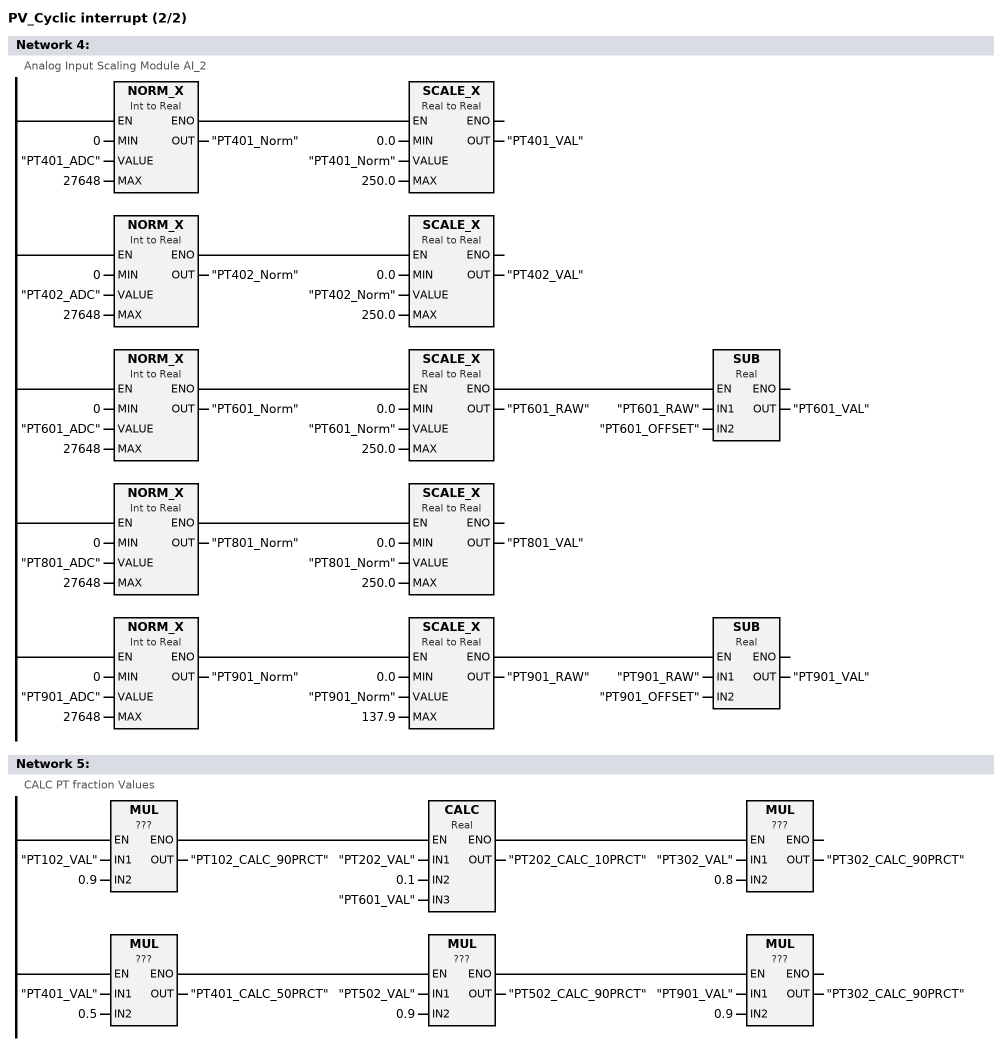
   RUNG wire#powerrail
      { S7_Templates := "[SrcType := Int, DestType := Real]" } Normalize(min := 0, value := "PT401_ADC", max := 27648, out => "PT401_Norm")
      { S7_Templates := "[SrcType := Real, DestType := Real]" } Scale(min := 0.0, value := "PT401_Norm", max := 250.0, out => "PT401_VAL")
   END_RUNG
   RUNG wire#powerrail
      { S7_Templates := "[SrcType := Int, DestType := Real]" } Normalize(min := 0, value := "PT402_ADC", max := 27648, out => "PT402_Norm")
      { S7_Templates := "[SrcType := Real, DestType := Real]" } Scale(min := 0.0, value := "PT402_Norm", max := 250.0, out => "PT402_VAL")
   END_RUNG
   RUNG wire#powerrail
      { S7_Templates := "[SrcType := Int, DestType := Real]" } Normalize(min := 0, value := "PT601_ADC", max := 27648, out => "PT601_Norm")
      { S7_Templates := "[SrcType := Real, DestType := Real]" } Scale(min := 0.0, value := "PT601_Norm", max := 250.0, out => "PT601_RAW")
      { S7_Templates := "SrcType := Real" } Sub(in1 := "PT601_RAW", in2 := "PT601_OFFSET", out => "PT601_VAL")
   END_RUNG
   RUNG wire#powerrail
      { S7_Templates := "[SrcType := Int, DestType := Real]" } Normalize(min := 0, value := "PT801_ADC", max := 27648, out => "PT801_Norm")
      { S7_Templates := "[SrcType := Real, DestType := Real]" } Scale(min := 0.0, value := "PT801_Norm", max := 250.0, out => "PT801_VAL")
   END_RUNG
   RUNG wire#powerrail
      { S7_Templates := "[SrcType := Int, DestType := Real]" } Normalize(min := 0, value := "PT901_ADC", max := 27648, out => "PT901_Norm")
      { S7_Templates := "[SrcType := Real, DestType := Real]" } Scale(min := 0.0, value := "PT901_Norm", max := 137.9, out => "PT901_RAW")
      { S7_Templates := "SrcType := Real" } Sub(in1 := "PT901_RAW", in2 := "PT901_OFFSET", out => "PT901_VAL")
   END_RUNG
   // the same network as SCL:
   "PT401_Norm" := NORM_X(MIN := 0, VALUE := "PT401_ADC", MAX := 27648);
   "PT401_VAL" := SCALE_X(MIN := 0.0, VALUE := "PT401_Norm", MAX := 250.0);
   "PT402_Norm" := NORM_X(MIN := 0, VALUE := "PT402_ADC", MAX := 27648);
   "PT402_VAL" := SCALE_X(MIN := 0.0, VALUE := "PT402_Norm", MAX := 250.0);
   "PT601_Norm" := NORM_X(MIN := 0, VALUE := "PT601_ADC", MAX := 27648);
   "PT601_RAW" := SCALE_X(MIN := 0.0, VALUE := "PT601_Norm", MAX := 250.0);
   "PT601_VAL" := "PT601_RAW" - "PT601_OFFSET";
   "PT801_Norm" := NORM_X(MIN := 0, VALUE := "PT801_ADC", MAX := 27648);
   "PT801_VAL" := SCALE_X(MIN := 0.0, VALUE := "PT801_Norm", MAX := 250.0);
   "PT901_Norm" := NORM_X(MIN := 0, VALUE := "PT901_ADC", MAX := 27648);
   "PT901_RAW" := SCALE_X(MIN := 0.0, VALUE := "PT901_Norm", MAX := 137.9);
   "PT901_VAL" := "PT901_RAW" - "PT901_OFFSET";
END_REGION

REGION Network 5
   // CALC PT fraction Values
   "PT102_CALC_90PRCT" := "PT102_VAL" * 0.9;
   CALC(in1 := "PT202_VAL", in2 := 0.1, in3 := "PT601_VAL", out => "PT202_CALC_10PRCT");
   "PT302_CALC_90PRCT" := "PT302_VAL" * 0.8;
   "PT401_CALC_50PRCT" := "PT401_VAL" * 0.5;
   "PT502_CALC_90PRCT" := "PT502_VAL" * 0.9;
   "PT302_CALC_90PRCT" := "PT901_VAL" * 0.9;
END_REGION
END_ORGANIZATION_BLOCK

ORGANIZATION_BLOCK "Startup"   // OB100, LAD, Startup
TITLE = "Complete Restart"
{ S7_Optimized_Access := 'FALSE' }
VERSION : 0.1
BEGIN

REGION Network 1
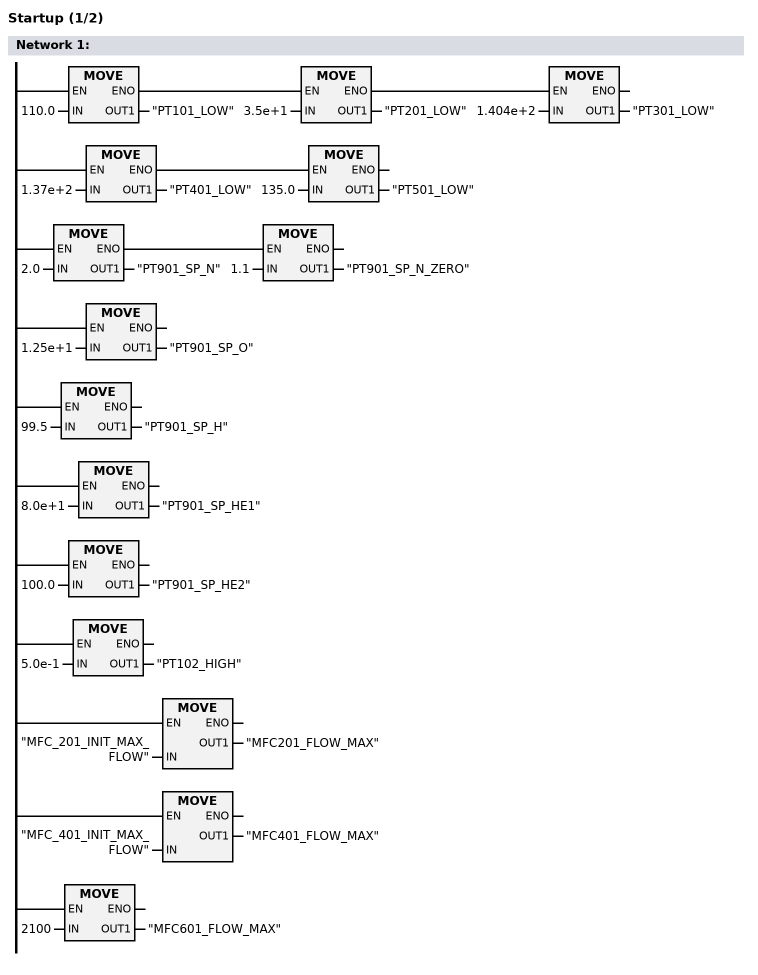
   RUNG wire#powerrail
      { S7_GenerateENO := "TRUE" } Move(in := 110.0, out1 => "PT101_LOW")
      { S7_GenerateENO := "TRUE" } Move(in := 3.5e+1, out1 => "PT201_LOW")
      { S7_GenerateENO := "TRUE" } Move(in := 1.404e+2, out1 => "PT301_LOW")
   END_RUNG
   RUNG wire#powerrail
      { S7_GenerateENO := "TRUE" } Move(in := 1.37e+2, out1 => "PT401_LOW")
      { S7_GenerateENO := "TRUE" } Move(in := 135.0, out1 => "PT501_LOW")
   END_RUNG
   RUNG wire#powerrail
      { S7_GenerateENO := "TRUE" } Move(in := 2.0, out1 => "PT901_SP_N")
      { S7_GenerateENO := "TRUE" } Move(in := 1.1, out1 => "PT901_SP_N_ZERO")
   END_RUNG
   RUNG wire#powerrail
      { S7_GenerateENO := "TRUE" } Move(in := 1.25e+1, out1 => "PT901_SP_O")
   END_RUNG
   RUNG wire#powerrail
      { S7_GenerateENO := "TRUE" } Move(in := 99.5, out1 => "PT901_SP_H")
   END_RUNG
   RUNG wire#powerrail
      { S7_GenerateENO := "TRUE" } Move(in := 8.0e+1, out1 => "PT901_SP_HE1")
   END_RUNG
   RUNG wire#powerrail
      { S7_GenerateENO := "TRUE" } Move(in := 100.0, out1 => "PT901_SP_HE2")
   END_RUNG
   RUNG wire#powerrail
      { S7_GenerateENO := "TRUE" } Move(in := 5.0e-1, out1 => "PT102_HIGH")
   END_RUNG
   RUNG wire#powerrail
      { S7_GenerateENO := "TRUE" } Move(in := "MFC_201_INIT_MAX_FLOW", out1 => "MFC201_FLOW_MAX")
   END_RUNG
   RUNG wire#powerrail
      { S7_GenerateENO := "TRUE" } Move(in := "MFC_401_INIT_MAX_FLOW", out1 => "MFC401_FLOW_MAX")
   END_RUNG
   RUNG wire#powerrail
      { S7_GenerateENO := "TRUE" } Move(in := 2100, out1 => "MFC601_FLOW_MAX")
   END_RUNG
   // the same network as SCL:
   // ENO of a box is taken as its EN; it also drops when the box reports an error
   "PT101_LOW" := 110.0;
   "PT201_LOW" := 3.5e+1;
   "PT301_LOW" := 1.404e+2;
   "PT401_LOW" := 1.37e+2;
   "PT501_LOW" := 135.0;
   "PT901_SP_N" := 2.0;
   "PT901_SP_N_ZERO" := 1.1;
   "PT901_SP_O" := 1.25e+1;
   "PT901_SP_H" := 99.5;
   "PT901_SP_HE1" := 8.0e+1;
   "PT901_SP_HE2" := 100.0;
   "PT102_HIGH" := 5.0e-1;
   "MFC201_FLOW_MAX" := "MFC_201_INIT_MAX_FLOW";
   "MFC401_FLOW_MAX" := "MFC_401_INIT_MAX_FLOW";
   "MFC601_FLOW_MAX" := 2100;
END_REGION

REGION Network 2
   // MODBUS MASTER Init
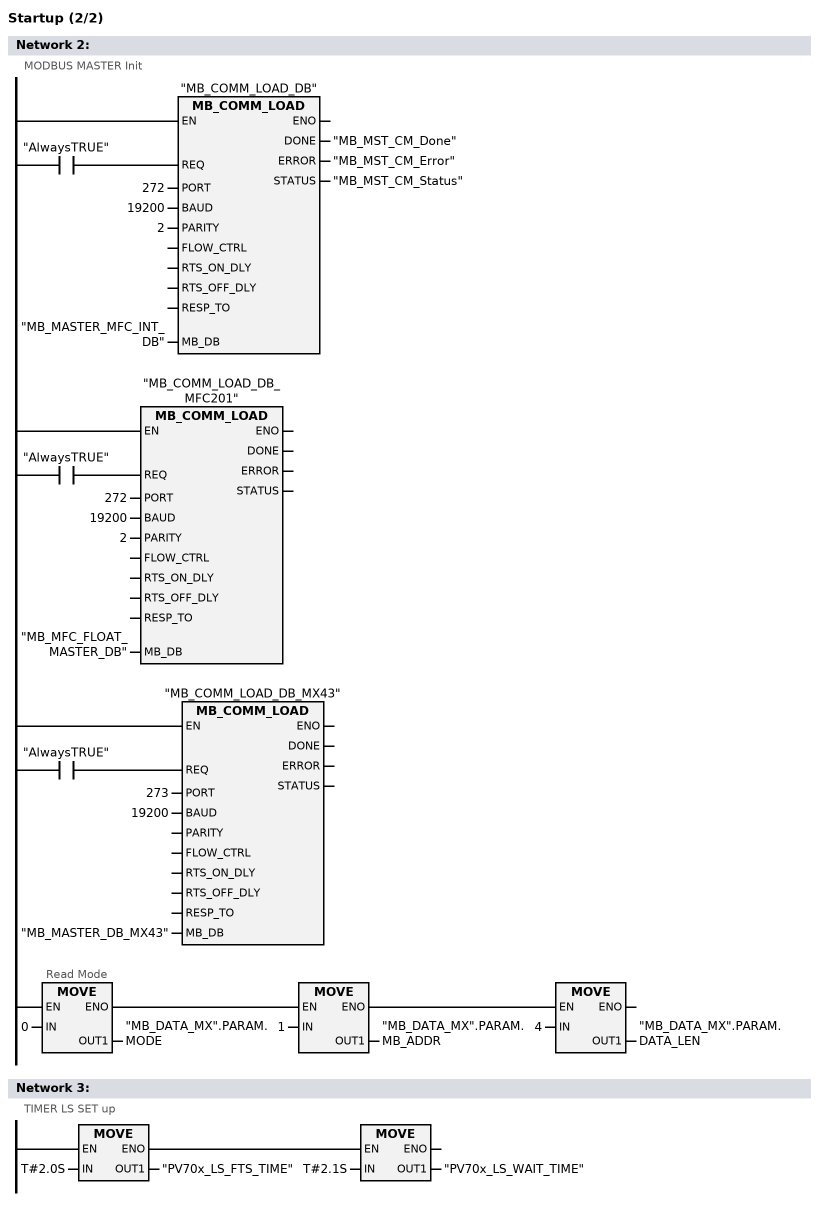
   "MB_COMM_LOAD_DB"(REQ := "AlwaysTRUE",   // MB_COMM_LOAD
                     PORT := 272,
                     BAUD := 19200,
                     PARITY := 2,
                     MB_DB := "MB_MASTER_MFC_INT_DB",
                     DONE => "MB_MST_CM_Done",
                     ERROR => "MB_MST_CM_Error",
                     STATUS => "MB_MST_CM_Status");
   "MB_COMM_LOAD_DB_MFC201"(REQ := "AlwaysTRUE",   // MB_COMM_LOAD
                           PORT := 272,
                           BAUD := 19200,
                           PARITY := 2,
                           MB_DB := "MB_MFC_FLOAT_MASTER_DB");
   "MB_COMM_LOAD_DB_MX43"(REQ := "AlwaysTRUE", PORT := 273, BAUD := 19200, MB_DB := "MB_MASTER_DB_MX43");   // MB_COMM_LOAD
   "MB_DATA_MX".PARAM.MODE := 0;   // Read Mode
   "MB_DATA_MX".PARAM.MB_ADDR := 1;
   "MB_DATA_MX".PARAM.DATA_LEN := 4;
END_REGION

REGION Network 3
   // TIMER LS SET up
   RUNG wire#powerrail
      Move(in := T#2.0S, out1 => "PV70x_LS_FTS_TIME")
      Move(in := T#2.1S, out1 => "PV70x_LS_WAIT_TIME")
   END_RUNG
   // the same network as SCL:
   "PV70x_LS_FTS_TIME" := T#2.0S;
   "PV70x_LS_WAIT_TIME" := T#2.1S;
END_REGION
END_ORGANIZATION_BLOCK